REGION Network 198
   RUNG wire#powerrail
      Contact( "Carrier_69_Status.7" )
      wire#w1
      Coil( "EMS".Carrier[69].CommFlt )
   END_RUNG
   RUNG wire#powerrail
      Contact( "C69_Heartbeat_On_Timer".Q )
   END_RUNG wire#w1
   RUNG wire#powerrail
      Contact( "C69_Heartbeat_Off_Timer".Q )
   END_RUNG wire#w1
   // the same network as SCL:
   "EMS".Carrier[69].CommFlt := "Carrier_69_Status.7" OR "C69_Heartbeat_On_Timer".Q OR "C69_Heartbeat_Off_Timer".Q;
END_REGION

REGION Network 199
   RUNG wire#powerrail
      Contact( "EMS".Carrier[69].CommFlt )
      JumpCoil( C69_Comm_Fault )
   END_RUNG
   // the same network as SCL:
   IF "EMS".Carrier[69].CommFlt THEN GOTO C69_Comm_Fault; END_IF;
END_REGION

REGION Network 200
   RUNG wire#powerrail
      { S7_Templates := "SrcType := Word" } NE_Contact(in1 := "Carrier_69_CarrierNumber", in2 := 0)
      Move(in := "Carrier_69_CarrierNumber", out1 => "EMS".Carrier[69].SDC_IN.CarrierNumber)
   END_RUNG
   // the same network as SCL:
   IF "Carrier_69_CarrierNumber" <> 0 THEN
       "EMS".Carrier[69].SDC_IN.CarrierNumber := "Carrier_69_CarrierNumber";
   END_IF;
END_REGION

REGION Network 201
   RUNG wire#powerrail
      { S7_Templates := "SrcType := DWord" } NE_Contact(in1 := "Carrier_69_CarrierPosition", in2 := 0)
      Move(in := "Carrier_69_CarrierPosition", out1 => "EMS".Carrier[69].SDC_IN.CarrierPosition)
   END_RUNG
   // the same network as SCL:
   IF "Carrier_69_CarrierPosition" <> 0 THEN
       "EMS".Carrier[69].SDC_IN.CarrierPosition := "Carrier_69_CarrierPosition";
   END_IF;
END_REGION

REGION Network 202
   RUNG wire#powerrail
      Move(in := "Carrier_69_ActualSpeed", out1 => "EMS".Carrier[69].SDC_IN.ActualSpeed)
   END_RUNG
   // the same network as SCL:
   "EMS".Carrier[69].SDC_IN.ActualSpeed := "Carrier_69_ActualSpeed";
END_REGION

REGION Network 203
   RUNG wire#powerrail
      Move(in := "Carrier_69_G120DControlWord", out1 => "DB402_SDC_CARRIER_DRIVE_DATA".Drive_Data.CARRIER[69].Drive_Control)
      Move(in := "Carrier_69_G120DStatusWord", out1 => "DB402_SDC_CARRIER_DRIVE_DATA".Drive_Data.CARRIER[69].Drive_Status)
   END_RUNG
   // the same network as SCL:
   "DB402_SDC_CARRIER_DRIVE_DATA".Drive_Data.CARRIER[69].Drive_Control := "Carrier_69_G120DControlWord";
   "DB402_SDC_CARRIER_DRIVE_DATA".Drive_Data.CARRIER[69].Drive_Status := "Carrier_69_G120DStatusWord";
END_REGION

REGION Network 204
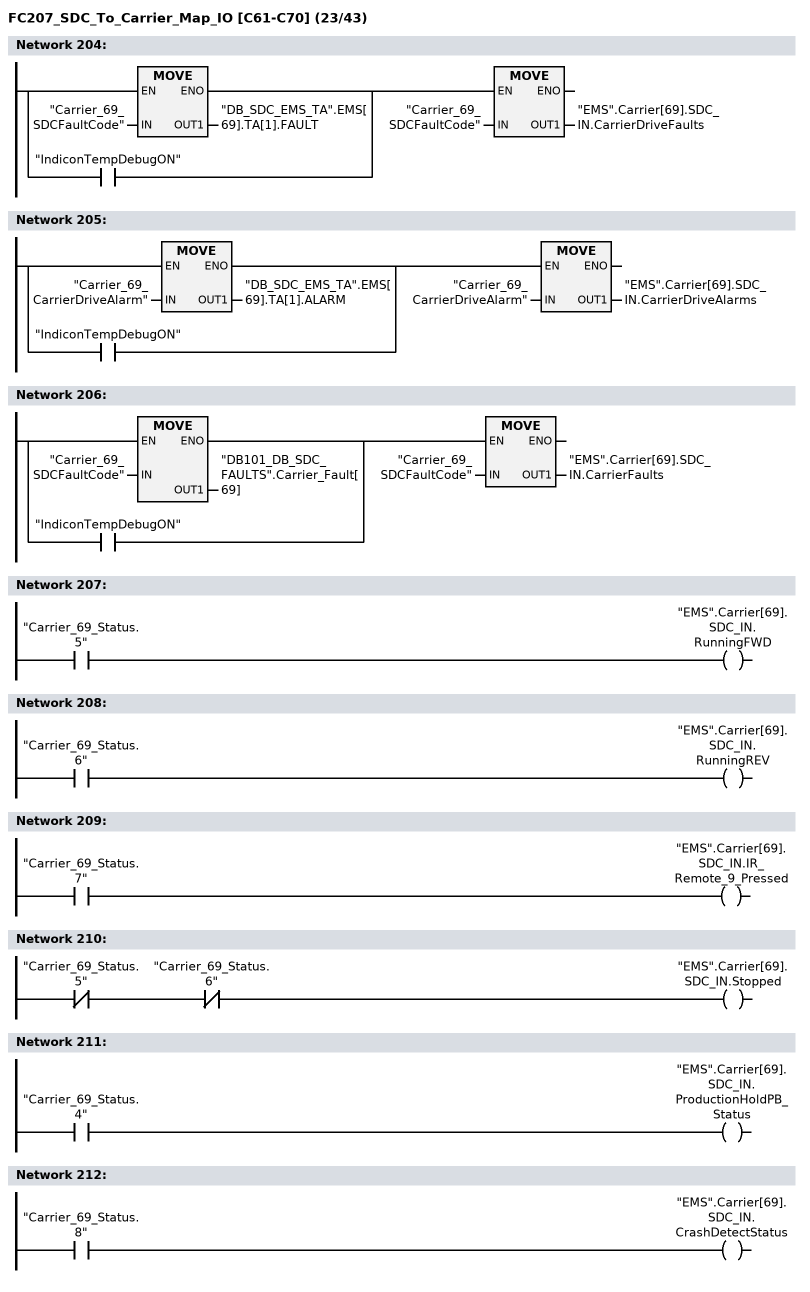
   RUNG wire#powerrail
      Move(in := "Carrier_69_SDCFaultCode", out1 => "DB_SDC_EMS_TA".EMS[69].TA[1].FAULT)
      wire#w1
      Move(in := "Carrier_69_SDCFaultCode", out1 => "EMS".Carrier[69].SDC_IN.CarrierDriveFaults)
   END_RUNG
   RUNG wire#powerrail
      Contact( "IndiconTempDebugON" )
   END_RUNG wire#w1
   // the same network as SCL:
   "DB_SDC_EMS_TA".EMS[69].TA[1].FAULT := "Carrier_69_SDCFaultCode";
   IF TRUE OR "IndiconTempDebugON" THEN
       "EMS".Carrier[69].SDC_IN.CarrierDriveFaults := "Carrier_69_SDCFaultCode";
   END_IF;
END_REGION

REGION Network 205
   RUNG wire#powerrail
      Move(in := "Carrier_69_CarrierDriveAlarm", out1 => "DB_SDC_EMS_TA".EMS[69].TA[1].ALARM)
      wire#w1
      Move(in := "Carrier_69_CarrierDriveAlarm", out1 => "EMS".Carrier[69].SDC_IN.CarrierDriveAlarms)
   END_RUNG
   RUNG wire#powerrail
      Contact( "IndiconTempDebugON" )
   END_RUNG wire#w1
   // the same network as SCL:
   "DB_SDC_EMS_TA".EMS[69].TA[1].ALARM := "Carrier_69_CarrierDriveAlarm";
   IF TRUE OR "IndiconTempDebugON" THEN
       "EMS".Carrier[69].SDC_IN.CarrierDriveAlarms := "Carrier_69_CarrierDriveAlarm";
   END_IF;
END_REGION

REGION Network 206
   RUNG wire#powerrail
      Move(in := "Carrier_69_SDCFaultCode", out1 => "DB101_DB_SDC_FAULTS".Carrier_Fault[69])
      wire#w1
      Move(in := "Carrier_69_SDCFaultCode", out1 => "EMS".Carrier[69].SDC_IN.CarrierFaults)
   END_RUNG
   RUNG wire#powerrail
      Contact( "IndiconTempDebugON" )
   END_RUNG wire#w1
   // the same network as SCL:
   "DB101_DB_SDC_FAULTS".Carrier_Fault[69] := "Carrier_69_SDCFaultCode";
   IF TRUE OR "IndiconTempDebugON" THEN
       "EMS".Carrier[69].SDC_IN.CarrierFaults := "Carrier_69_SDCFaultCode";
   END_IF;
END_REGION

REGION Network 207
   RUNG wire#powerrail
      Contact( "Carrier_69_Status.5" )
      Coil( "EMS".Carrier[69].SDC_IN.RunningFWD )
   END_RUNG
   // the same network as SCL:
   "EMS".Carrier[69].SDC_IN.RunningFWD := "Carrier_69_Status.5";
END_REGION

REGION Network 208
   RUNG wire#powerrail
      Contact( "Carrier_69_Status.6" )
      Coil( "EMS".Carrier[69].SDC_IN.RunningREV )
   END_RUNG
   // the same network as SCL:
   "EMS".Carrier[69].SDC_IN.RunningREV := "Carrier_69_Status.6";
END_REGION

REGION Network 209
   RUNG wire#powerrail
      Contact( "Carrier_69_Status.7" )
      Coil( "EMS".Carrier[69].SDC_IN.IR_Remote_9_Pressed )
   END_RUNG
   // the same network as SCL:
   "EMS".Carrier[69].SDC_IN.IR_Remote_9_Pressed := "Carrier_69_Status.7";
END_REGION

REGION Network 210
   RUNG wire#powerrail
      I_Contact( "Carrier_69_Status.5" )
      I_Contact( "Carrier_69_Status.6" )
      Coil( "EMS".Carrier[69].SDC_IN.Stopped )
   END_RUNG
   // the same network as SCL:
   "EMS".Carrier[69].SDC_IN.Stopped := NOT "Carrier_69_Status.5" AND NOT "Carrier_69_Status.6";
END_REGION

REGION Network 211
   RUNG wire#powerrail
      Contact( "Carrier_69_Status.4" )
      Coil( "EMS".Carrier[69].SDC_IN.ProductionHoldPB_Status )
   END_RUNG
   // the same network as SCL:
   "EMS".Carrier[69].SDC_IN.ProductionHoldPB_Status := "Carrier_69_Status.4";
END_REGION

REGION Network 212
   RUNG wire#powerrail
      Contact( "Carrier_69_Status.8" )
      Coil( "EMS".Carrier[69].SDC_IN.CrashDetectStatus )
   END_RUNG
   // the same network as SCL:
   "EMS".Carrier[69].SDC_IN.CrashDetectStatus := "Carrier_69_Status.8";
END_REGION

REGION Network 213
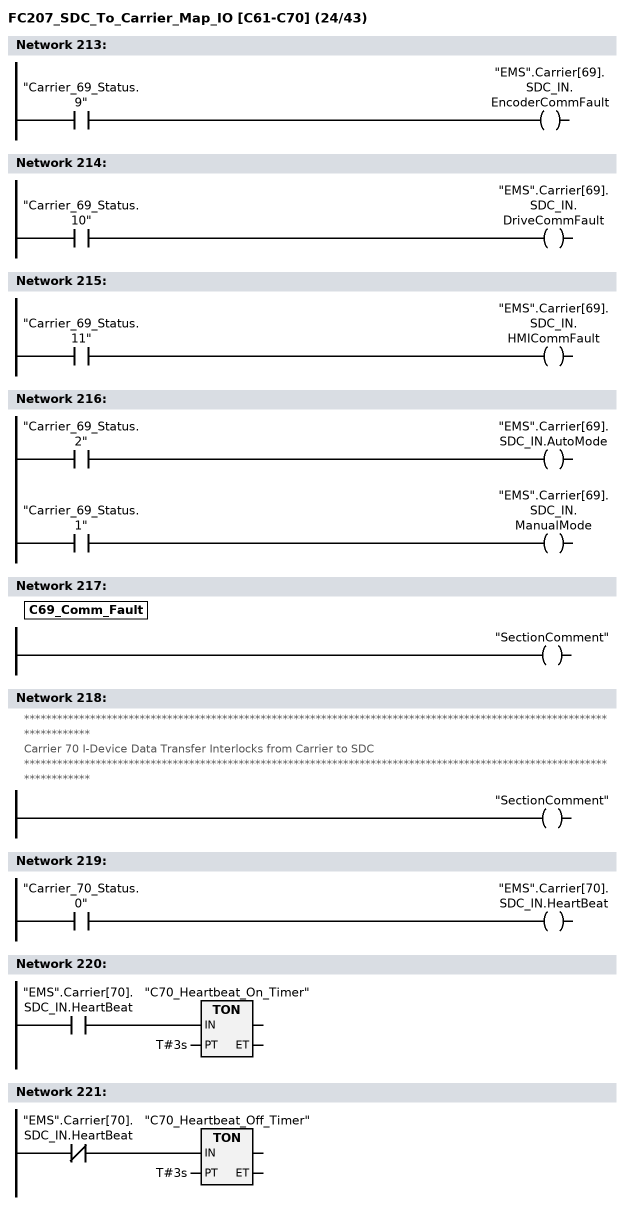
   RUNG wire#powerrail
      Contact( "Carrier_69_Status.9" )
      Coil( "EMS".Carrier[69].SDC_IN.EncoderCommFault )
   END_RUNG
   // the same network as SCL:
   "EMS".Carrier[69].SDC_IN.EncoderCommFault := "Carrier_69_Status.9";
END_REGION

REGION Network 214
   RUNG wire#powerrail
      Contact( "Carrier_69_Status.10" )
      Coil( "EMS".Carrier[69].SDC_IN.DriveCommFault )
   END_RUNG
   // the same network as SCL:
   "EMS".Carrier[69].SDC_IN.DriveCommFault := "Carrier_69_Status.10";
END_REGION

REGION Network 215
   RUNG wire#powerrail
      Contact( "Carrier_69_Status.11" )
      Coil( "EMS".Carrier[69].SDC_IN.HMICommFault )
   END_RUNG
   // the same network as SCL:
   "EMS".Carrier[69].SDC_IN.HMICommFault := "Carrier_69_Status.11";
END_REGION

REGION Network 216
   RUNG wire#powerrail
      Contact( "Carrier_69_Status.2" )
      Coil( "EMS".Carrier[69].SDC_IN.AutoMode )
   END_RUNG
   RUNG wire#powerrail
      Contact( "Carrier_69_Status.1" )
      Coil( "EMS".Carrier[69].SDC_IN.ManualMode )
   END_RUNG
   // the same network as SCL:
   "EMS".Carrier[69].SDC_IN.AutoMode := "Carrier_69_Status.2";
   "EMS".Carrier[69].SDC_IN.ManualMode := "Carrier_69_Status.1";
END_REGION

REGION Network 217
   Label( C69_Comm_Fault )
   RUNG wire#powerrail
      Coil( "SectionComment" )
   END_RUNG
   // the same network as SCL:
   C69_Comm_Fault:
   "SectionComment" := TRUE;
END_REGION

REGION Network 218
   // **********************************************************************************************************************
   // 
   // Carrier 70 I-Device Data Transfer Interlocks from Carrier to SDC
   // 
   // **********************************************************************************************************************
   RUNG wire#powerrail
      Coil( "SectionComment" )
   END_RUNG
   // the same network as SCL:
   "SectionComment" := TRUE;
END_REGION

REGION Network 219
   RUNG wire#powerrail
      Contact( "Carrier_70_Status.0" )
      Coil( "EMS".Carrier[70].SDC_IN.HeartBeat )
   END_RUNG
   // the same network as SCL:
   "EMS".Carrier[70].SDC_IN.HeartBeat := "Carrier_70_Status.0";
END_REGION

REGION Network 220
   "C70_Heartbeat_On_Timer".TON(IN := "EMS".Carrier[70].SDC_IN.HeartBeat, PT := T#3s);
END_REGION

REGION Network 221
   "C70_Heartbeat_Off_Timer".TON(IN := NOT "EMS".Carrier[70].SDC_IN.HeartBeat, PT := T#3s);
END_REGION

REGION Network 222
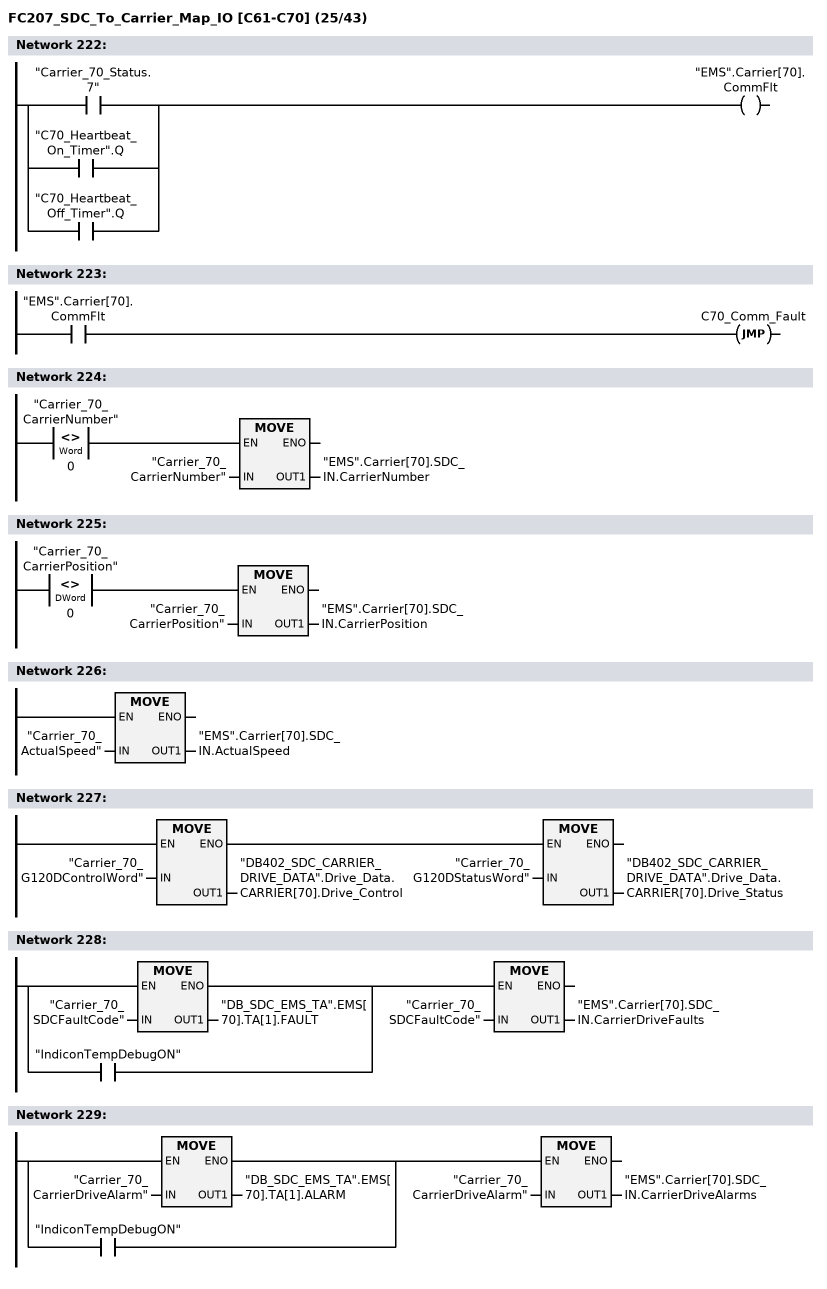
   RUNG wire#powerrail
      Contact( "Carrier_70_Status.7" )
      wire#w1
      Coil( "EMS".Carrier[70].CommFlt )
   END_RUNG
   RUNG wire#powerrail
      Contact( "C70_Heartbeat_On_Timer".Q )
   END_RUNG wire#w1
   RUNG wire#powerrail
      Contact( "C70_Heartbeat_Off_Timer".Q )
   END_RUNG wire#w1
   // the same network as SCL:
   "EMS".Carrier[70].CommFlt := "Carrier_70_Status.7" OR "C70_Heartbeat_On_Timer".Q OR "C70_Heartbeat_Off_Timer".Q;
END_REGION

REGION Network 223
   RUNG wire#powerrail
      Contact( "EMS".Carrier[70].CommFlt )
      JumpCoil( C70_Comm_Fault )
   END_RUNG
   // the same network as SCL:
   IF "EMS".Carrier[70].CommFlt THEN GOTO C70_Comm_Fault; END_IF;
END_REGION

REGION Network 224
   RUNG wire#powerrail
      { S7_Templates := "SrcType := Word" } NE_Contact(in1 := "Carrier_70_CarrierNumber", in2 := 0)
      Move(in := "Carrier_70_CarrierNumber", out1 => "EMS".Carrier[70].SDC_IN.CarrierNumber)
   END_RUNG
   // the same network as SCL:
   IF "Carrier_70_CarrierNumber" <> 0 THEN
       "EMS".Carrier[70].SDC_IN.CarrierNumber := "Carrier_70_CarrierNumber";
   END_IF;
END_REGION

REGION Network 225
   RUNG wire#powerrail
      { S7_Templates := "SrcType := DWord" } NE_Contact(in1 := "Carrier_70_CarrierPosition", in2 := 0)
      Move(in := "Carrier_70_CarrierPosition", out1 => "EMS".Carrier[70].SDC_IN.CarrierPosition)
   END_RUNG
   // the same network as SCL:
   IF "Carrier_70_CarrierPosition" <> 0 THEN
       "EMS".Carrier[70].SDC_IN.CarrierPosition := "Carrier_70_CarrierPosition";
   END_IF;
END_REGION

REGION Network 226
   RUNG wire#powerrail
      Move(in := "Carrier_70_ActualSpeed", out1 => "EMS".Carrier[70].SDC_IN.ActualSpeed)
   END_RUNG
   // the same network as SCL:
   "EMS".Carrier[70].SDC_IN.ActualSpeed := "Carrier_70_ActualSpeed";
END_REGION

REGION Network 227
   RUNG wire#powerrail
      Move(in := "Carrier_70_G120DControlWord", out1 => "DB402_SDC_CARRIER_DRIVE_DATA".Drive_Data.CARRIER[70].Drive_Control)
      Move(in := "Carrier_70_G120DStatusWord", out1 => "DB402_SDC_CARRIER_DRIVE_DATA".Drive_Data.CARRIER[70].Drive_Status)
   END_RUNG
   // the same network as SCL:
   "DB402_SDC_CARRIER_DRIVE_DATA".Drive_Data.CARRIER[70].Drive_Control := "Carrier_70_G120DControlWord";
   "DB402_SDC_CARRIER_DRIVE_DATA".Drive_Data.CARRIER[70].Drive_Status := "Carrier_70_G120DStatusWord";
END_REGION

REGION Network 228
   RUNG wire#powerrail
      Move(in := "Carrier_70_SDCFaultCode", out1 => "DB_SDC_EMS_TA".EMS[70].TA[1].FAULT)
      wire#w1
      Move(in := "Carrier_70_SDCFaultCode", out1 => "EMS".Carrier[70].SDC_IN.CarrierDriveFaults)
   END_RUNG
   RUNG wire#powerrail
      Contact( "IndiconTempDebugON" )
   END_RUNG wire#w1
   // the same network as SCL:
   "DB_SDC_EMS_TA".EMS[70].TA[1].FAULT := "Carrier_70_SDCFaultCode";
   IF TRUE OR "IndiconTempDebugON" THEN
       "EMS".Carrier[70].SDC_IN.CarrierDriveFaults := "Carrier_70_SDCFaultCode";
   END_IF;
END_REGION

REGION Network 229
   RUNG wire#powerrail
      Move(in := "Carrier_70_CarrierDriveAlarm", out1 => "DB_SDC_EMS_TA".EMS[70].TA[1].ALARM)
      wire#w1
      Move(in := "Carrier_70_CarrierDriveAlarm", out1 => "EMS".Carrier[70].SDC_IN.CarrierDriveAlarms)
   END_RUNG
   RUNG wire#powerrail
      Contact( "IndiconTempDebugON" )
   END_RUNG wire#w1
   // the same network as SCL:
   "DB_SDC_EMS_TA".EMS[70].TA[1].ALARM := "Carrier_70_CarrierDriveAlarm";
   IF TRUE OR "IndiconTempDebugON" THEN
       "EMS".Carrier[70].SDC_IN.CarrierDriveAlarms := "Carrier_70_CarrierDriveAlarm";
   END_IF;
END_REGION

REGION Network 230
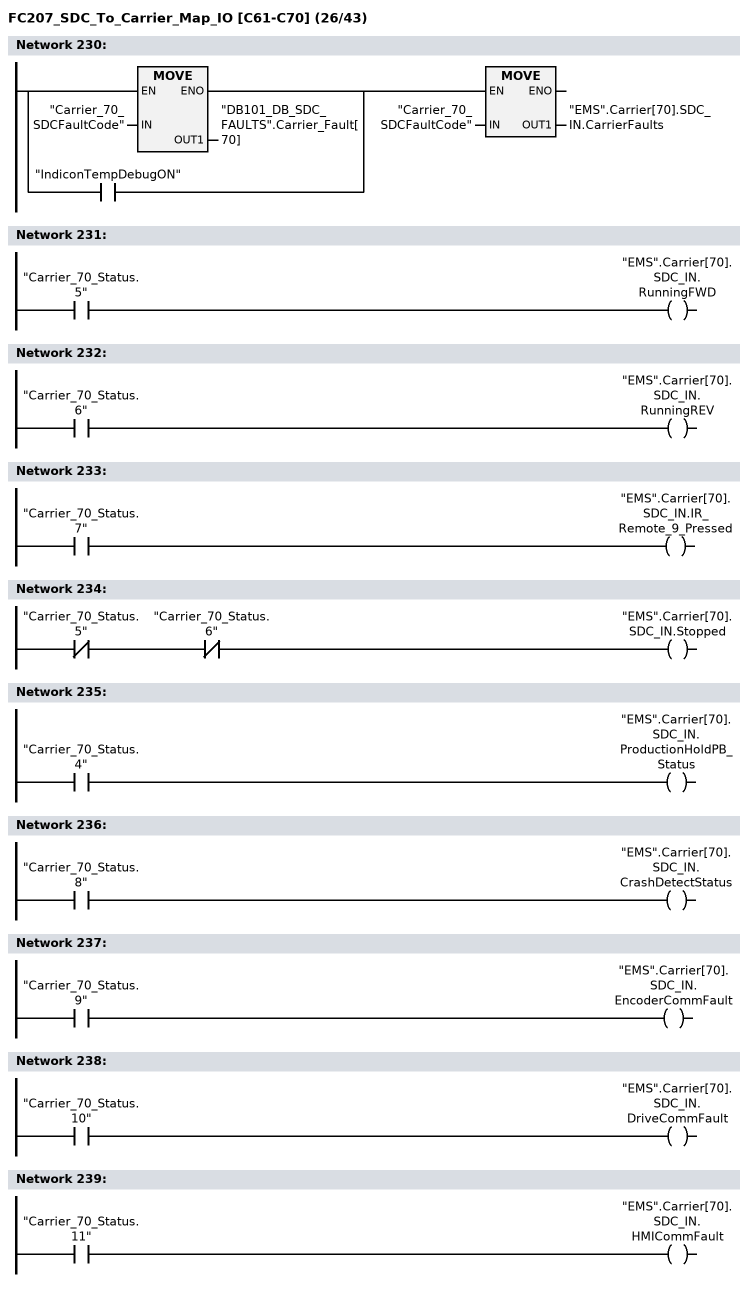
   RUNG wire#powerrail
      Move(in := "Carrier_70_SDCFaultCode", out1 => "DB101_DB_SDC_FAULTS".Carrier_Fault[70])
      wire#w1
      Move(in := "Carrier_70_SDCFaultCode", out1 => "EMS".Carrier[70].SDC_IN.CarrierFaults)
   END_RUNG
   RUNG wire#powerrail
      Contact( "IndiconTempDebugON" )
   END_RUNG wire#w1
   // the same network as SCL:
   "DB101_DB_SDC_FAULTS".Carrier_Fault[70] := "Carrier_70_SDCFaultCode";
   IF TRUE OR "IndiconTempDebugON" THEN
       "EMS".Carrier[70].SDC_IN.CarrierFaults := "Carrier_70_SDCFaultCode";
   END_IF;
END_REGION

REGION Network 231
   RUNG wire#powerrail
      Contact( "Carrier_70_Status.5" )
      Coil( "EMS".Carrier[70].SDC_IN.RunningFWD )
   END_RUNG
   // the same network as SCL:
   "EMS".Carrier[70].SDC_IN.RunningFWD := "Carrier_70_Status.5";
END_REGION

REGION Network 232
   RUNG wire#powerrail
      Contact( "Carrier_70_Status.6" )
      Coil( "EMS".Carrier[70].SDC_IN.RunningREV )
   END_RUNG
   // the same network as SCL:
   "EMS".Carrier[70].SDC_IN.RunningREV := "Carrier_70_Status.6";
END_REGION

REGION Network 233
   RUNG wire#powerrail
      Contact( "Carrier_70_Status.7" )
      Coil( "EMS".Carrier[70].SDC_IN.IR_Remote_9_Pressed )
   END_RUNG
   // the same network as SCL:
   "EMS".Carrier[70].SDC_IN.IR_Remote_9_Pressed := "Carrier_70_Status.7";
END_REGION

REGION Network 234
   RUNG wire#powerrail
      I_Contact( "Carrier_70_Status.5" )
      I_Contact( "Carrier_70_Status.6" )
      Coil( "EMS".Carrier[70].SDC_IN.Stopped )
   END_RUNG
   // the same network as SCL:
   "EMS".Carrier[70].SDC_IN.Stopped := NOT "Carrier_70_Status.5" AND NOT "Carrier_70_Status.6";
END_REGION

REGION Network 235
   RUNG wire#powerrail
      Contact( "Carrier_70_Status.4" )
      Coil( "EMS".Carrier[70].SDC_IN.ProductionHoldPB_Status )
   END_RUNG
   // the same network as SCL:
   "EMS".Carrier[70].SDC_IN.ProductionHoldPB_Status := "Carrier_70_Status.4";
END_REGION

REGION Network 236
   RUNG wire#powerrail
      Contact( "Carrier_70_Status.8" )
      Coil( "EMS".Carrier[70].SDC_IN.CrashDetectStatus )
   END_RUNG
   // the same network as SCL:
   "EMS".Carrier[70].SDC_IN.CrashDetectStatus := "Carrier_70_Status.8";
END_REGION

REGION Network 237
   RUNG wire#powerrail
      Contact( "Carrier_70_Status.9" )
      Coil( "EMS".Carrier[70].SDC_IN.EncoderCommFault )
   END_RUNG
   // the same network as SCL:
   "EMS".Carrier[70].SDC_IN.EncoderCommFault := "Carrier_70_Status.9";
END_REGION

REGION Network 238
   RUNG wire#powerrail
      Contact( "Carrier_70_Status.10" )
      Coil( "EMS".Carrier[70].SDC_IN.DriveCommFault )
   END_RUNG
   // the same network as SCL:
   "EMS".Carrier[70].SDC_IN.DriveCommFault := "Carrier_70_Status.10";
END_REGION

REGION Network 239
   RUNG wire#powerrail
      Contact( "Carrier_70_Status.11" )
      Coil( "EMS".Carrier[70].SDC_IN.HMICommFault )
   END_RUNG
   // the same network as SCL:
   "EMS".Carrier[70].SDC_IN.HMICommFault := "Carrier_70_Status.11";
END_REGION

REGION Network 240
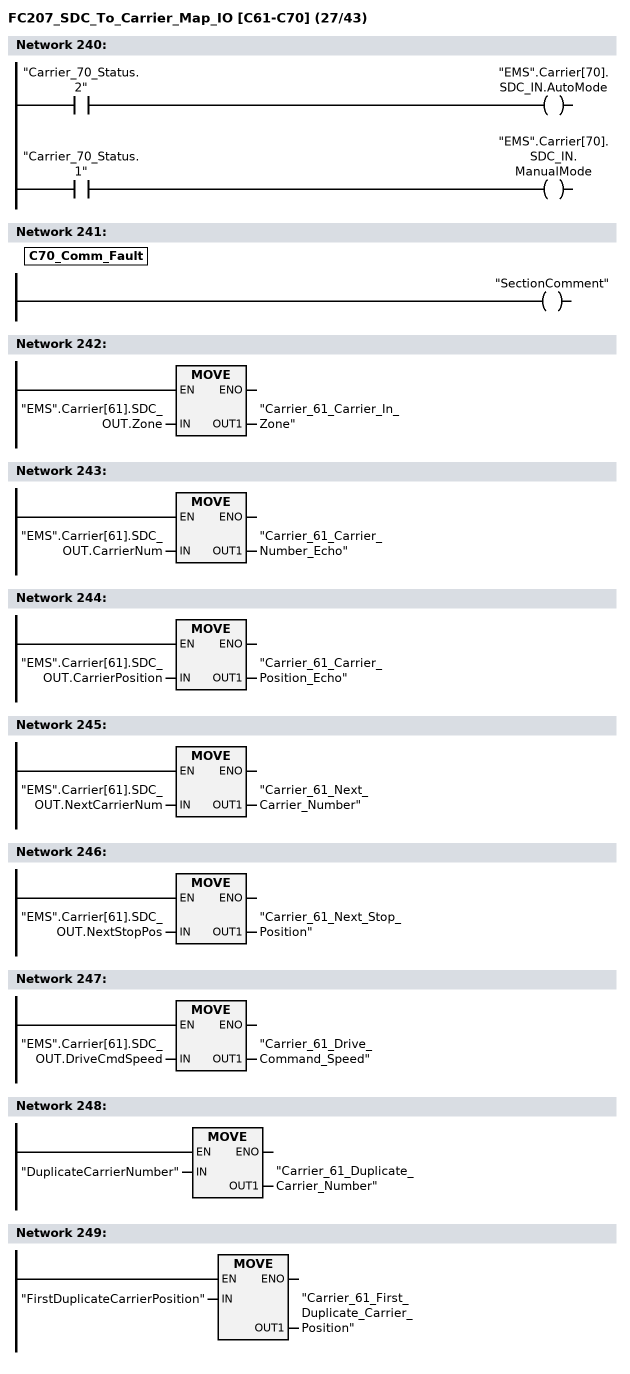
   RUNG wire#powerrail
      Contact( "Carrier_70_Status.2" )
      Coil( "EMS".Carrier[70].SDC_IN.AutoMode )
   END_RUNG
   RUNG wire#powerrail
      Contact( "Carrier_70_Status.1" )
      Coil( "EMS".Carrier[70].SDC_IN.ManualMode )
   END_RUNG
   // the same network as SCL:
   "EMS".Carrier[70].SDC_IN.AutoMode := "Carrier_70_Status.2";
   "EMS".Carrier[70].SDC_IN.ManualMode := "Carrier_70_Status.1";
END_REGION

REGION Network 241
   Label( C70_Comm_Fault )
   RUNG wire#powerrail
      Coil( "SectionComment" )
   END_RUNG
   // the same network as SCL:
   C70_Comm_Fault:
   "SectionComment" := TRUE;
END_REGION

REGION Network 242
   RUNG wire#powerrail
      Move(in := "EMS".Carrier[61].SDC_OUT.Zone, out1 => "Carrier_61_Carrier_In_Zone")
   END_RUNG
   // the same network as SCL:
   "Carrier_61_Carrier_In_Zone" := "EMS".Carrier[61].SDC_OUT.Zone;
END_REGION

REGION Network 243
   RUNG wire#powerrail
      Move(in := "EMS".Carrier[61].SDC_OUT.CarrierNum, out1 => "Carrier_61_Carrier_Number_Echo")
   END_RUNG
   // the same network as SCL:
   "Carrier_61_Carrier_Number_Echo" := "EMS".Carrier[61].SDC_OUT.CarrierNum;
END_REGION

REGION Network 244
   RUNG wire#powerrail
      Move(in := "EMS".Carrier[61].SDC_OUT.CarrierPosition, out1 => "Carrier_61_Carrier_Position_Echo")
   END_RUNG
   // the same network as SCL:
   "Carrier_61_Carrier_Position_Echo" := "EMS".Carrier[61].SDC_OUT.CarrierPosition;
END_REGION

REGION Network 245
   RUNG wire#powerrail
      Move(in := "EMS".Carrier[61].SDC_OUT.NextCarrierNum, out1 => "Carrier_61_Next_Carrier_Number")
   END_RUNG
   // the same network as SCL:
   "Carrier_61_Next_Carrier_Number" := "EMS".Carrier[61].SDC_OUT.NextCarrierNum;
END_REGION

REGION Network 246
   RUNG wire#powerrail
      Move(in := "EMS".Carrier[61].SDC_OUT.NextStopPos, out1 => "Carrier_61_Next_Stop_Position")
   END_RUNG
   // the same network as SCL:
   "Carrier_61_Next_Stop_Position" := "EMS".Carrier[61].SDC_OUT.NextStopPos;
END_REGION

REGION Network 247
   RUNG wire#powerrail
      Move(in := "EMS".Carrier[61].SDC_OUT.DriveCmdSpeed, out1 => "Carrier_61_Drive_Command_Speed")
   END_RUNG
   // the same network as SCL:
   "Carrier_61_Drive_Command_Speed" := "EMS".Carrier[61].SDC_OUT.DriveCmdSpeed;
END_REGION

REGION Network 248
   RUNG wire#powerrail
      Move(in := "DuplicateCarrierNumber", out1 => "Carrier_61_Duplicate_Carrier_Number")
   END_RUNG
   // the same network as SCL:
   "Carrier_61_Duplicate_Carrier_Number" := "DuplicateCarrierNumber";
END_REGION

REGION Network 249
   RUNG wire#powerrail
      Move(in := "FirstDuplicateCarrierPosition", out1 => "Carrier_61_First_Duplicate_Carrier_Position")
   END_RUNG
   // the same network as SCL:
   "Carrier_61_First_Duplicate_Carrier_Position" := "FirstDuplicateCarrierPosition";
END_REGION

REGION Network 250
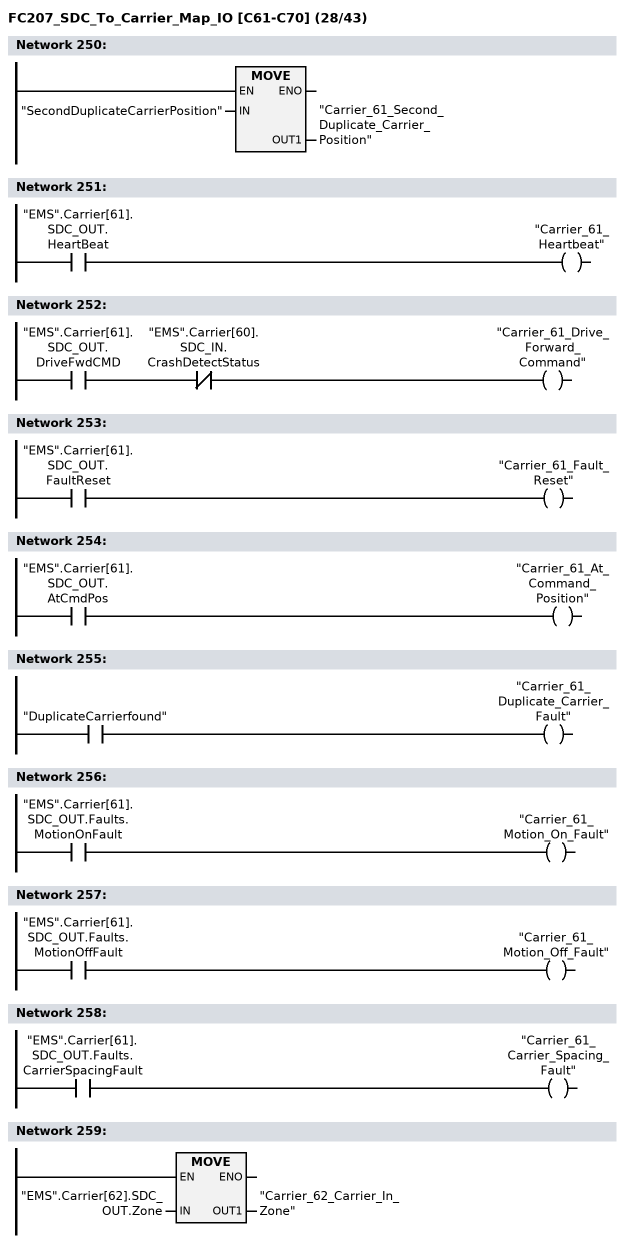
   RUNG wire#powerrail
      Move(in := "SecondDuplicateCarrierPosition", out1 => "Carrier_61_Second_Duplicate_Carrier_Position")
   END_RUNG
   // the same network as SCL:
   "Carrier_61_Second_Duplicate_Carrier_Position" := "SecondDuplicateCarrierPosition";
END_REGION

REGION Network 251
   RUNG wire#powerrail
      Contact( "EMS".Carrier[61].SDC_OUT.HeartBeat )
      Coil( "Carrier_61_Heartbeat" )
   END_RUNG
   // the same network as SCL:
   "Carrier_61_Heartbeat" := "EMS".Carrier[61].SDC_OUT.HeartBeat;
END_REGION

REGION Network 252
   RUNG wire#powerrail
      Contact( "EMS".Carrier[61].SDC_OUT.DriveFwdCMD )
      I_Contact( "EMS".Carrier[60].SDC_IN.CrashDetectStatus )
      Coil( "Carrier_61_Drive_Forward_Command" )
   END_RUNG
   // the same network as SCL:
   "Carrier_61_Drive_Forward_Command" := "EMS".Carrier[61].SDC_OUT.DriveFwdCMD AND NOT "EMS".Carrier[60].SDC_IN.CrashDetectStatus;
END_REGION

REGION Network 253
   RUNG wire#powerrail
      Contact( "EMS".Carrier[61].SDC_OUT.FaultReset )
      Coil( "Carrier_61_Fault_Reset" )
   END_RUNG
   // the same network as SCL:
   "Carrier_61_Fault_Reset" := "EMS".Carrier[61].SDC_OUT.FaultReset;
END_REGION

REGION Network 254
   RUNG wire#powerrail
      Contact( "EMS".Carrier[61].SDC_OUT.AtCmdPos )
      Coil( "Carrier_61_At_Command_Position" )
   END_RUNG
   // the same network as SCL:
   "Carrier_61_At_Command_Position" := "EMS".Carrier[61].SDC_OUT.AtCmdPos;
END_REGION

REGION Network 255
   RUNG wire#powerrail
      Contact( "DuplicateCarrierfound" )
      Coil( "Carrier_61_Duplicate_Carrier_Fault" )
   END_RUNG
   // the same network as SCL:
   "Carrier_61_Duplicate_Carrier_Fault" := "DuplicateCarrierfound";
END_REGION

REGION Network 256
   RUNG wire#powerrail
      Contact( "EMS".Carrier[61].SDC_OUT.Faults.MotionOnFault )
      Coil( "Carrier_61_Motion_On_Fault" )
   END_RUNG
   // the same network as SCL:
   "Carrier_61_Motion_On_Fault" := "EMS".Carrier[61].SDC_OUT.Faults.MotionOnFault;
END_REGION

REGION Network 257
   RUNG wire#powerrail
      Contact( "EMS".Carrier[61].SDC_OUT.Faults.MotionOffFault )
      Coil( "Carrier_61_Motion_Off_Fault" )
   END_RUNG
   // the same network as SCL:
   "Carrier_61_Motion_Off_Fault" := "EMS".Carrier[61].SDC_OUT.Faults.MotionOffFault;
END_REGION

REGION Network 258
   RUNG wire#powerrail
      Contact( "EMS".Carrier[61].SDC_OUT.Faults.CarrierSpacingFault )
      Coil( "Carrier_61_Carrier_Spacing_Fault" )
   END_RUNG
   // the same network as SCL:
   "Carrier_61_Carrier_Spacing_Fault" := "EMS".Carrier[61].SDC_OUT.Faults.CarrierSpacingFault;
END_REGION

REGION Network 259
   RUNG wire#powerrail
      Move(in := "EMS".Carrier[62].SDC_OUT.Zone, out1 => "Carrier_62_Carrier_In_Zone")
   END_RUNG
   // the same network as SCL:
   "Carrier_62_Carrier_In_Zone" := "EMS".Carrier[62].SDC_OUT.Zone;
END_REGION

REGION Network 260
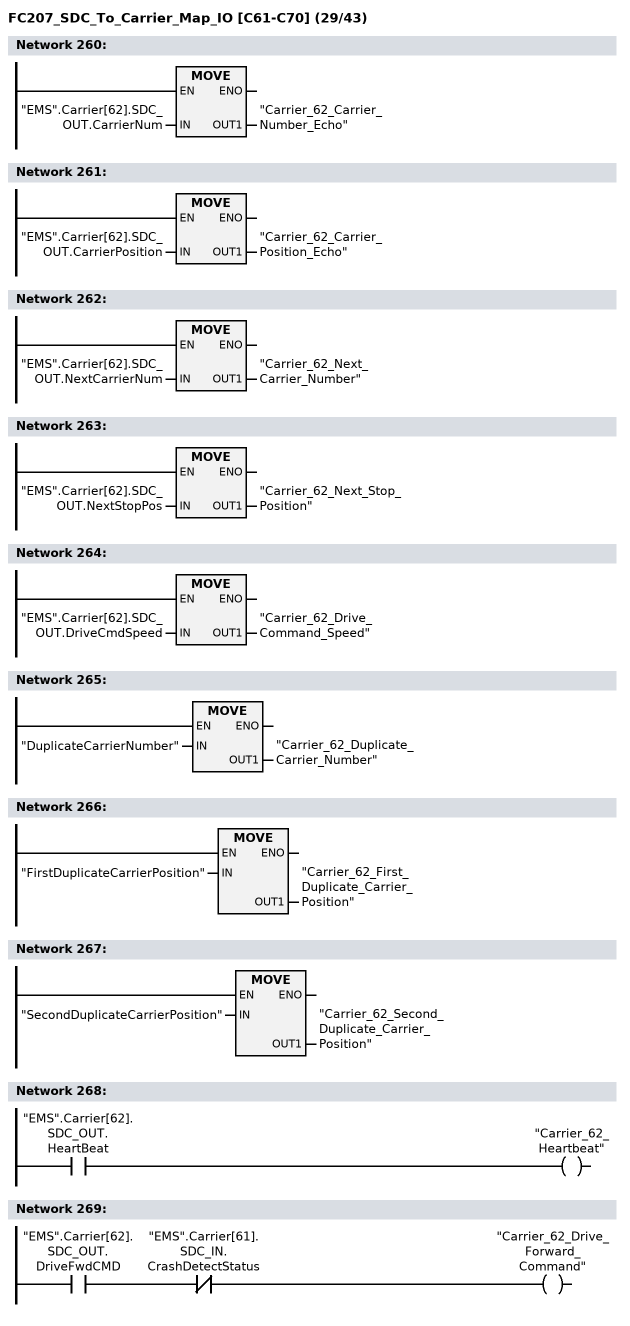
   RUNG wire#powerrail
      Move(in := "EMS".Carrier[62].SDC_OUT.CarrierNum, out1 => "Carrier_62_Carrier_Number_Echo")
   END_RUNG
   // the same network as SCL:
   "Carrier_62_Carrier_Number_Echo" := "EMS".Carrier[62].SDC_OUT.CarrierNum;
END_REGION

REGION Network 261
   RUNG wire#powerrail
      Move(in := "EMS".Carrier[62].SDC_OUT.CarrierPosition, out1 => "Carrier_62_Carrier_Position_Echo")
   END_RUNG
   // the same network as SCL:
   "Carrier_62_Carrier_Position_Echo" := "EMS".Carrier[62].SDC_OUT.CarrierPosition;
END_REGION

REGION Network 262
   RUNG wire#powerrail
      Move(in := "EMS".Carrier[62].SDC_OUT.NextCarrierNum, out1 => "Carrier_62_Next_Carrier_Number")
   END_RUNG
   // the same network as SCL:
   "Carrier_62_Next_Carrier_Number" := "EMS".Carrier[62].SDC_OUT.NextCarrierNum;
END_REGION

REGION Network 263
   RUNG wire#powerrail
      Move(in := "EMS".Carrier[62].SDC_OUT.NextStopPos, out1 => "Carrier_62_Next_Stop_Position")
   END_RUNG
   // the same network as SCL:
   "Carrier_62_Next_Stop_Position" := "EMS".Carrier[62].SDC_OUT.NextStopPos;
END_REGION

REGION Network 264
   RUNG wire#powerrail
      Move(in := "EMS".Carrier[62].SDC_OUT.DriveCmdSpeed, out1 => "Carrier_62_Drive_Command_Speed")
   END_RUNG
   // the same network as SCL:
   "Carrier_62_Drive_Command_Speed" := "EMS".Carrier[62].SDC_OUT.DriveCmdSpeed;
END_REGION

REGION Network 265
   RUNG wire#powerrail
      Move(in := "DuplicateCarrierNumber", out1 => "Carrier_62_Duplicate_Carrier_Number")
   END_RUNG
   // the same network as SCL:
   "Carrier_62_Duplicate_Carrier_Number" := "DuplicateCarrierNumber";
END_REGION

REGION Network 266
   RUNG wire#powerrail
      Move(in := "FirstDuplicateCarrierPosition", out1 => "Carrier_62_First_Duplicate_Carrier_Position")
   END_RUNG
   // the same network as SCL:
   "Carrier_62_First_Duplicate_Carrier_Position" := "FirstDuplicateCarrierPosition";
END_REGION

REGION Network 267
   RUNG wire#powerrail
      Move(in := "SecondDuplicateCarrierPosition", out1 => "Carrier_62_Second_Duplicate_Carrier_Position")
   END_RUNG
   // the same network as SCL:
   "Carrier_62_Second_Duplicate_Carrier_Position" := "SecondDuplicateCarrierPosition";
END_REGION

REGION Network 268
   RUNG wire#powerrail
      Contact( "EMS".Carrier[62].SDC_OUT.HeartBeat )
      Coil( "Carrier_62_Heartbeat" )
   END_RUNG
   // the same network as SCL:
   "Carrier_62_Heartbeat" := "EMS".Carrier[62].SDC_OUT.HeartBeat;
END_REGION

REGION Network 269
   RUNG wire#powerrail
      Contact( "EMS".Carrier[62].SDC_OUT.DriveFwdCMD )
      I_Contact( "EMS".Carrier[61].SDC_IN.CrashDetectStatus )
      Coil( "Carrier_62_Drive_Forward_Command" )
   END_RUNG
   // the same network as SCL:
   "Carrier_62_Drive_Forward_Command" := "EMS".Carrier[62].SDC_OUT.DriveFwdCMD AND NOT "EMS".Carrier[61].SDC_IN.CrashDetectStatus;
END_REGION

REGION Network 270
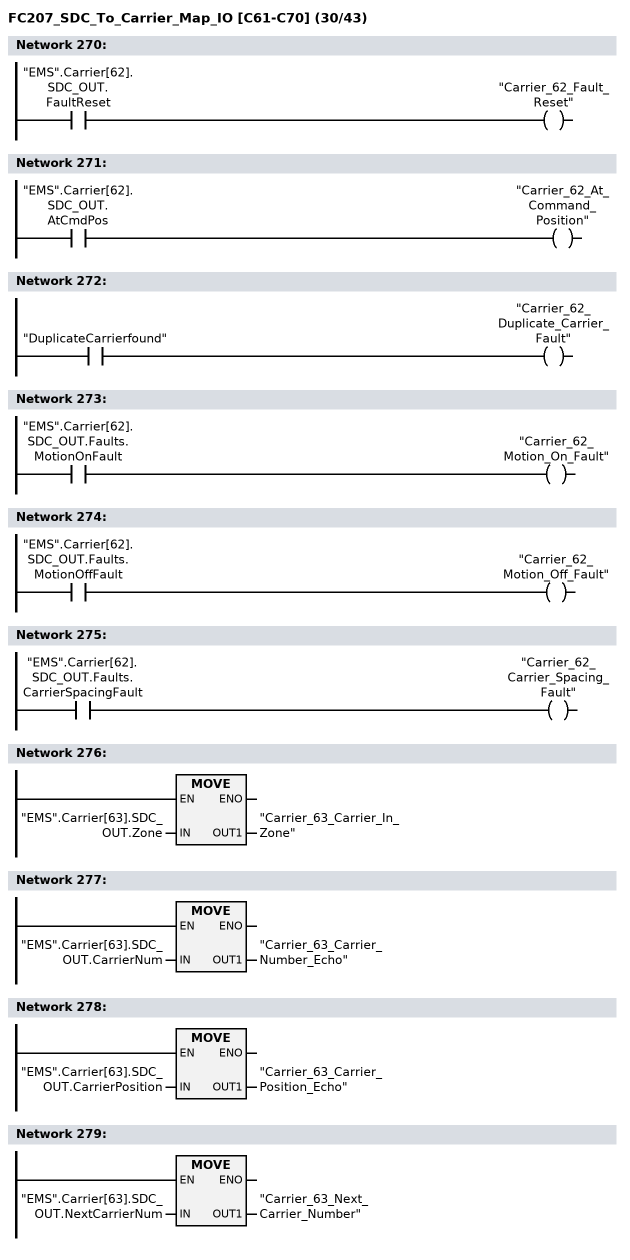
   RUNG wire#powerrail
      Contact( "EMS".Carrier[62].SDC_OUT.FaultReset )
      Coil( "Carrier_62_Fault_Reset" )
   END_RUNG
   // the same network as SCL:
   "Carrier_62_Fault_Reset" := "EMS".Carrier[62].SDC_OUT.FaultReset;
END_REGION

REGION Network 271
   RUNG wire#powerrail
      Contact( "EMS".Carrier[62].SDC_OUT.AtCmdPos )
      Coil( "Carrier_62_At_Command_Position" )
   END_RUNG
   // the same network as SCL:
   "Carrier_62_At_Command_Position" := "EMS".Carrier[62].SDC_OUT.AtCmdPos;
END_REGION

REGION Network 272
   RUNG wire#powerrail
      Contact( "DuplicateCarrierfound" )
      Coil( "Carrier_62_Duplicate_Carrier_Fault" )
   END_RUNG
   // the same network as SCL:
   "Carrier_62_Duplicate_Carrier_Fault" := "DuplicateCarrierfound";
END_REGION

REGION Network 273
   RUNG wire#powerrail
      Contact( "EMS".Carrier[62].SDC_OUT.Faults.MotionOnFault )
      Coil( "Carrier_62_Motion_On_Fault" )
   END_RUNG
   // the same network as SCL:
   "Carrier_62_Motion_On_Fault" := "EMS".Carrier[62].SDC_OUT.Faults.MotionOnFault;
END_REGION

REGION Network 274
   RUNG wire#powerrail
      Contact( "EMS".Carrier[62].SDC_OUT.Faults.MotionOffFault )
      Coil( "Carrier_62_Motion_Off_Fault" )
   END_RUNG
   // the same network as SCL:
   "Carrier_62_Motion_Off_Fault" := "EMS".Carrier[62].SDC_OUT.Faults.MotionOffFault;
END_REGION

REGION Network 275
   RUNG wire#powerrail
      Contact( "EMS".Carrier[62].SDC_OUT.Faults.CarrierSpacingFault )
      Coil( "Carrier_62_Carrier_Spacing_Fault" )
   END_RUNG
   // the same network as SCL:
   "Carrier_62_Carrier_Spacing_Fault" := "EMS".Carrier[62].SDC_OUT.Faults.CarrierSpacingFault;
END_REGION

REGION Network 276
   RUNG wire#powerrail
      Move(in := "EMS".Carrier[63].SDC_OUT.Zone, out1 => "Carrier_63_Carrier_In_Zone")
   END_RUNG
   // the same network as SCL:
   "Carrier_63_Carrier_In_Zone" := "EMS".Carrier[63].SDC_OUT.Zone;
END_REGION

REGION Network 277
   RUNG wire#powerrail
      Move(in := "EMS".Carrier[63].SDC_OUT.CarrierNum, out1 => "Carrier_63_Carrier_Number_Echo")
   END_RUNG
   // the same network as SCL:
   "Carrier_63_Carrier_Number_Echo" := "EMS".Carrier[63].SDC_OUT.CarrierNum;
END_REGION

REGION Network 278
   RUNG wire#powerrail
      Move(in := "EMS".Carrier[63].SDC_OUT.CarrierPosition, out1 => "Carrier_63_Carrier_Position_Echo")
   END_RUNG
   // the same network as SCL:
   "Carrier_63_Carrier_Position_Echo" := "EMS".Carrier[63].SDC_OUT.CarrierPosition;
END_REGION

REGION Network 279
   RUNG wire#powerrail
      Move(in := "EMS".Carrier[63].SDC_OUT.NextCarrierNum, out1 => "Carrier_63_Next_Carrier_Number")
   END_RUNG
   // the same network as SCL:
   "Carrier_63_Next_Carrier_Number" := "EMS".Carrier[63].SDC_OUT.NextCarrierNum;
END_REGION

REGION Network 280
